// TIA Portal project "Project_ModbusTCPIP" (V15.1)

(* hardware
DEVICE "S7-1200 station_1"  S7-1200 Station
   slot 0: "Rack_0"  S7-1200 Rack  Rack  V1.0
   slot 1: "S71200_Station1"  CPU 1212FC DC/DC/DC  6ES7 212-1AF40-0XB0  V4.2
DEVICE "S7-1200 station_2"  S7-1200 Station
   slot 0: "Rack_0"  S7-1200 Rack  Rack  V1.0
   slot 1: "S71200_Station2"  CPU 1217C DC/DC/DC  6ES7 217-1AG40-0XB0  V4.2
DEVICE "HMI_1"  TP900 Comfort
   slot 0: "HMI_1"  TP900 Comfort  6AV2 124-0JC01-0AX0  15.1.0.0
   slot 1: "HMI_RT_1"  TP900 Comfort  6AV2 124-0JC01-0AX0  15.1.0.0
   slot 5: "HMI_1.IE_CP_1"  PROFINET Interface  15.0.1.0
      slot 1: "PROFINET Interface_1"  PROFINET Interface
         slot 1: "Port_1"  Port
         slot 2: "Port_2"  Port
   slot 7: "HMI_1.MPI/DP_CP_1"  MPI/DP Interface  15.0.1.0
*)

// ===== PLC "S71200_Station1"  CPU 1212FC DC/DC/DC =====

VAR_GLOBAL   // PLC tag table "Default tag table"
   "M_DISCONNECT" AT %M0.0 : Bool;
END_VAR

DATA_BLOCK "dbConfig"   // DB2
{ S7_Optimized_Access := 'TRUE' }
VERSION : 0.1
   VAR
      CONNECT : TCON_IP_v4;
   END_VAR
BEGIN
   CONNECT.InterfaceId := 1;
   CONNECT.ID := 16#001;
   CONNECT.ConnectionType := 16#0B;
   CONNECT.ActiveEstablished := FALSE;
   CONNECT.RemoteAddress.ADDR[1] := 16#C0;
   CONNECT.RemoteAddress.ADDR[2] := 16#A8;
   CONNECT.RemoteAddress.ADDR[3] := 16#0B;
   CONNECT.RemoteAddress.ADDR[4] := 16#32;
   CONNECT.RemotePort := 0;
   CONNECT.LocalPort := 5900;
END_DATA_BLOCK

DATA_BLOCK "dbMB_HOLD_REG"   // DB3
{ S7_Optimized_Access := 'FALSE' }
VERSION : 0.1
   VAR
      r : Array[0..9] of Int;
   END_VAR
BEGIN
END_DATA_BLOCK

ORGANIZATION_BLOCK "Main"   // OB1, LAD, ProgramCycle
TITLE = "Main Program Sweep (Cycle)"
{ S7_Optimized_Access := 'TRUE' }
VERSION : 0.1
   VAR_INPUT
      Initial_Call : Bool;   // Initial call of this OB
      Remanence : Bool;   // =True, if remanent data are available
   END_VAR
BEGIN

REGION Network 1
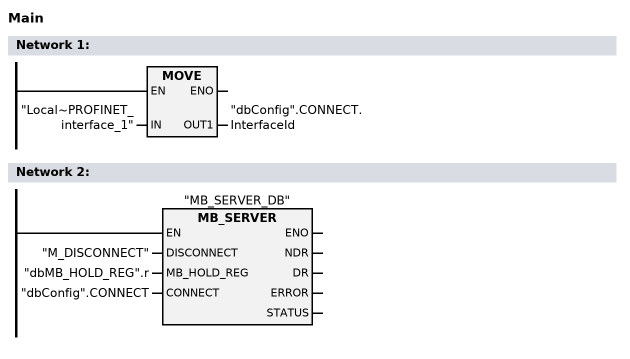
   RUNG wire#powerrail
      Move(in := "Local~PROFINET_interface_1", out1 => "dbConfig".CONNECT.InterfaceId)
   END_RUNG
   // the same network as SCL:
   "dbConfig".CONNECT.InterfaceId := "Local~PROFINET_interface_1";
END_REGION

REGION Network 2
   "MB_SERVER_DB"(DISCONNECT := "M_DISCONNECT", MB_HOLD_REG := "dbMB_HOLD_REG".r, CONNECT := "dbConfig".CONNECT);   // MB_SERVER
END_REGION
END_ORGANIZATION_BLOCK

// ===== PLC "S71200_Station2"  CPU 1217C DC/DC/DC =====

VAR_GLOBAL   // PLC tag table "Default tag table"
   "M_DISCONNECT" AT %M0.0 : Bool;
END_VAR

DATA_BLOCK "dbConfig"   // DB2
{ S7_Optimized_Access := 'TRUE' }
VERSION : 0.1
   VAR
      CONNECT : TCON_IP_v4;
   END_VAR
BEGIN
   CONNECT.InterfaceId := 1;
   CONNECT.ID := 16#001;
   CONNECT.ConnectionType := 16#0B;
   CONNECT.ActiveEstablished := FALSE;
   CONNECT.RemoteAddress.ADDR[1] := 16#C0;
   CONNECT.RemoteAddress.ADDR[2] := 16#A8;
   CONNECT.RemoteAddress.ADDR[3] := 16#0B;
   CONNECT.RemoteAddress.ADDR[4] := 16#32;
   CONNECT.RemotePort := 0;
   CONNECT.LocalPort := 5900;
END_DATA_BLOCK

DATA_BLOCK "dbMB_HOLD_REG"   // DB3
{ S7_Optimized_Access := 'FALSE' }
VERSION : 0.1
   VAR
      r : Array[0..9] of Int;
      w : Array[0..9] of Int;
   END_VAR
BEGIN
END_DATA_BLOCK

ORGANIZATION_BLOCK "Main"   // OB1, LAD, ProgramCycle
TITLE = "Main Program Sweep (Cycle)"
{ S7_Optimized_Access := 'TRUE' }
VERSION : 0.1
   VAR_INPUT
      Initial_Call : Bool;   // Initial call of this OB
      Remanence : Bool;   // =True, if remanent data are available
   END_VAR
BEGIN

REGION Network 1
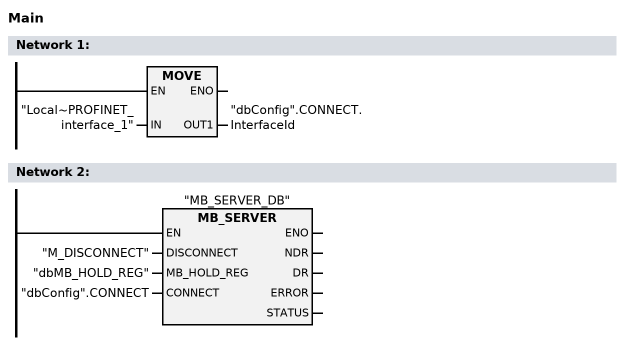
   RUNG wire#powerrail
      Move(in := "Local~PROFINET_interface_1", out1 => "dbConfig".CONNECT.InterfaceId)
   END_RUNG
   // the same network as SCL:
   "dbConfig".CONNECT.InterfaceId := "Local~PROFINET_interface_1";
END_REGION

REGION Network 2
   "MB_SERVER_DB"(DISCONNECT := "M_DISCONNECT", MB_HOLD_REG := "dbMB_HOLD_REG", CONNECT := "dbConfig".CONNECT);   // MB_SERVER
END_REGION
END_ORGANIZATION_BLOCK

(* ===== HMI "HMI_RT_1" =====
system functions are stored by id; their names below are inferred from use
connection "HMI_S71200_Station1": ETHERNET, S7_1200_OMS
connection "HMI_S71200_Station2": ETHERNET, S7_1200_OMS

HMI tags "Default tag table"
   "Tag_ScreenNumber" : UInt, internal

HMI tags "_S71200_Station1"
   "S71200_Station1_dbMB_HOLD_REG_r" : Array [0..9] of Int = PLC dbMB_HOLD_REG.r AT %DB3.DBX0.0, 1 s

HMI tags "_S71200_Station2"
   "S71200_Station2_dbMB_HOLD_REG_r" : Array [0..9] of Int = PLC dbMB_HOLD_REG.r AT %DB3.DBX0.0, 1 s
   "S71200_Station2_dbMB_HOLD_REG_w" : Array [0..9] of Int = PLC dbMB_HOLD_REG.w AT %DB3.DBX20.0, 1 s

screen "Root screen" 800x420, template "Template_1"
   on GenerateScreen: SetTag("Tag_ScreenNumber", 1)
   IOField "I/O field_1" at 130,66 size 96x32; FormatPattern s99999
      ProcessValue <- "[0]"
   IOField "I/O field_2" at 130,99 size 96x32; FormatPattern s99999
      ProcessValue <- "[1]"
   IOField "I/O field_3" at 130,133 size 96x32; FormatPattern s99999
      ProcessValue <- "[2]"
   IOField "I/O field_4" at 130,167 size 96x32; FormatPattern s99999
      ProcessValue <- "[3]"
   IOField "I/O field_5" at 130,201 size 96x32; FormatPattern s99999
      ProcessValue <- "[4]"
   IOField "I/O field_6" at 130,234 size 96x32; FormatPattern s99999
      ProcessValue <- "[5]"
   IOField "I/O field_7" at 130,268 size 96x32; FormatPattern s99999
      ProcessValue <- "[6]"
   IOField "I/O field_8" at 130,302 size 96x32; FormatPattern s99999
      ProcessValue <- "[7]"
   IOField "I/O field_9" at 130,336 size 96x32; FormatPattern s99999
      ProcessValue <- "[8]"
   IOField "I/O field_10" at 130,370 size 96x32; FormatPattern s99999
      ProcessValue <- "[9]"
   TextField "Text field_1" at 131,12 size 94x50; Text 'S71200 Station1'
   TextField "Text field_2" at 72,69 size 56x27; Text '0x00'
   TextField "Text field_3" at 72,102 size 56x27; Text '0x01'
   TextField "Text field_4" at 72,136 size 56x27; Text '0x02'
   TextField "Text field_5" at 72,170 size 56x27; Text '0x03'
   TextField "Text field_6" at 72,204 size 56x27; Text '0x04'
   TextField "Text field_7" at 72,237 size 56x27; Text '0x05'
   TextField "Text field_8" at 72,271 size 56x27; Text '0x06'
   TextField "Text field_9" at 72,305 size 56x27; Text '0x07'
   TextField "Text field_10" at 72,339 size 56x27; Text '0x08'
   TextField "Text field_11" at 72,373 size 56x27; Text '0x09'
   Group "Group" at 72,12 size 154x390
   IOField "I/O field_11" at 335,66 size 96x32; FormatPattern s99999
      ProcessValue <- "[0]"
   IOField "I/O field_12" at 335,99 size 96x32; FormatPattern s99999
      ProcessValue <- "[1]"
   IOField "I/O field_13" at 335,133 size 96x32; FormatPattern s99999
      ProcessValue <- "[2]"
   IOField "I/O field_14" at 335,167 size 96x32; FormatPattern s99999
      ProcessValue <- "[3]"
   IOField "I/O field_15" at 335,201 size 96x32; FormatPattern s99999
      ProcessValue <- "[4]"
   IOField "I/O field_16" at 335,234 size 96x32; FormatPattern s99999
      ProcessValue <- "[5]"
   IOField "I/O field_17" at 335,268 size 96x32; FormatPattern s99999
      ProcessValue <- "[6]"
   IOField "I/O field_18" at 335,302 size 96x32; FormatPattern s99999
      ProcessValue <- "[7]"
   IOField "I/O field_19" at 335,336 size 96x32; FormatPattern s99999
      ProcessValue <- "[8]"
   IOField "I/O field_20" at 335,370 size 96x32; FormatPattern s99999
      ProcessValue <- "[9]"
   TextField "Text field_12" at 402,12 size 94x50; Text 'S71200 Station2'
   TextField "Text field_13" at 277,69 size 56x27; Text '0x00'
   TextField "Text field_14" at 277,102 size 56x27; Text '0x01'
   TextField "Text field_15" at 277,136 size 56x27; Text '0x02'
   TextField "Text field_16" at 277,170 size 56x27; Text '0x03'
   TextField "Text field_17" at 277,204 size 56x27; Text '0x04'
   TextField "Text field_18" at 277,237 size 56x27; Text '0x05'
   TextField "Text field_19" at 277,271 size 56x27; Text '0x06'
   TextField "Text field_20" at 277,305 size 56x27; Text '0x07'
   TextField "Text field_21" at 277,339 size 56x27; Text '0x08'
   TextField "Text field_22" at 277,373 size 56x27; Text '0x09'
   IOField "I/O field_21" at 511,66 size 96x32; FormatPattern s99999
      ProcessValue <- "[0]"
   IOField "I/O field_22" at 511,99 size 96x32; FormatPattern s99999
      ProcessValue <- "[1]"
   IOField "I/O field_23" at 511,133 size 96x32; FormatPattern s99999
      ProcessValue <- "[2]"
   IOField "I/O field_24" at 511,167 size 96x32; FormatPattern s99999
      ProcessValue <- "[3]"
   IOField "I/O field_25" at 511,201 size 96x32; FormatPattern s99999
      ProcessValue <- "[4]"
   IOField "I/O field_26" at 511,234 size 96x32; FormatPattern s99999
      ProcessValue <- "[5]"
   IOField "I/O field_27" at 511,268 size 96x32; FormatPattern s99999
      ProcessValue <- "[6]"
   IOField "I/O field_28" at 511,302 size 96x32; FormatPattern s99999
      ProcessValue <- "[7]"
   IOField "I/O field_29" at 511,336 size 96x32; FormatPattern s99999
      ProcessValue <- "[8]"
   IOField "I/O field_30" at 511,370 size 96x32; FormatPattern s99999
      ProcessValue <- "[9]"
   TextField "Text field_23" at 453,69 size 56x27; Text '0x00'
   TextField "Text field_24" at 453,102 size 56x27; Text '0x01'
   TextField "Text field_25" at 453,136 size 56x27; Text '0x02'
   TextField "Text field_26" at 453,170 size 56x27; Text '0x03'
   TextField "Text field_27" at 453,204 size 56x27; Text '0x04'
   TextField "Text field_28" at 453,237 size 56x27; Text '0x05'
   TextField "Text field_29" at 453,271 size 56x27; Text '0x06'
   TextField "Text field_30" at 453,305 size 56x27; Text '0x07'
   TextField "Text field_31" at 453,339 size 56x27; Text '0x08'
   TextField "Text field_32" at 453,373 size 56x27; Text '0x09'
*)